// TIA Portal project "RRI" (V15.1)

(* hardware
DEVICE "S7-1200 station_1"  S7-1200 Station
   slot 0: "Rack_0"  S7-1200 Rack  Rack  V1.0
   slot 1: "PLC_1"  CPU 1215C DC/DC/DC  6ES7 215-1AG40-0XB0  V4.3
   slot 2: "AI 4xRTD_1"  SM 1231 AI4 x RTD  6ES7 231-5PD32-0XB0  V2.0
   slot 3: "DI 16/DQ 16x24VDC_1"  6ES7 223-1BL32-0XB0  V2.0
DEVICE "GSD device_2"  GSD.Device.PN
   slot 0: "Rack"  Rack  V1.0
   slot 0: "clipx_M5"  0.25 ms, 6 slots  BMxx
      slot 0: "0.25 ms, 6 slots"  0.25 ms, 6 slots
      slot 1: "PN-IO"  PN-IO
         slot 1: "Port 1"  Port 1
         slot 2: "Port 2"  Port 2
   slot 1: "Max value_1"  Max value
      slot 0: "max value (REAL)"  max value (REAL)
   slot 2: "Min value_1"  Min value
      slot 0: "min value (REAL)"  min value (REAL)
DEVICE "GSD device_1"  GSD.Device.PN
   slot 0: "Rack"  Rack  V1.0
   slot 0: "ek9300-16"  EK9300 V2.3  EK9300  V1.00
      slot 0: "EK9300 V2.3_1"  EK9300 V2.3
      slot 1: "EK9300 V2.3"  EK9300 V2.3
         slot 1: "Port 1"  Port 1
         slot 2: "Port 2"  Port 2
   slot 1: "Standard"  Standard
   slot 1: "EL3068_1"  EL3068  EL3068
      slot 0: "ModuleAccessPoint"  ModuleAccessPoint
   slot 1: "Standard"  Standard
DEVICE "GSD device_3"  GSD.Device.PN
   slot 0: "Rack"  Rack  V1.0
   slot 0: "clipx_M1"  0.25 ms, 6 slots  BMxx
      slot 0: "0.25 ms, 6 slots"  0.25 ms, 6 slots
      slot 1: "PN-IO"  PN-IO
         slot 1: "Port 1"  Port 1
         slot 2: "Port 2"  Port 2
   slot 1: "Max value_1"  Max value
      slot 0: "max value (REAL)"  max value (REAL)
   slot 2: "Min value_1"  Min value
      slot 0: "min value (REAL)"  min value (REAL)
   slot 3: "Max value_2"  Max value
      slot 0: "max value (REAL)"  max value (REAL)
   slot 4: "Min value_2"  Min value
      slot 0: "min value (REAL)"  min value (REAL)
DEVICE "GSD device_4"  GSD.Device.PN
   slot 0: "Rack"  Rack  V1.0
   slot 0: "clipx_M2"  0.25 ms, 6 slots  BMxx
      slot 0: "0.25 ms, 6 slots"  0.25 ms, 6 slots
      slot 1: "PN-IO"  PN-IO
         slot 1: "Port 1"  Port 1
         slot 2: "Port 2"  Port 2
   slot 1: "Max value_1"  Max value
      slot 0: "max value (REAL)"  max value (REAL)
   slot 2: "Min value_1"  Min value
      slot 0: "min value (REAL)"  min value (REAL)
DEVICE "GSD device_5"  GSD.Device.PN
   slot 0: "Rack"  Rack  V1.0
   slot 0: "clipx_M3"  0.25 ms, 6 slots  BMxx
      slot 0: "0.25 ms, 6 slots"  0.25 ms, 6 slots
      slot 1: "PN-IO"  PN-IO
         slot 1: "Port 1"  Port 1
         slot 2: "Port 2"  Port 2
   slot 1: "Max value_1"  Max value
      slot 0: "max value (REAL)"  max value (REAL)
   slot 2: "Min value_1"  Min value
      slot 0: "min value (REAL)"  min value (REAL)
DEVICE "GSD device_6"  GSD.Device.PN
   slot 0: "Rack"  Rack  V1.0
   slot 0: "clipx_M4"  0.25 ms, 6 slots  BMxx
      slot 0: "0.25 ms, 6 slots"  0.25 ms, 6 slots
      slot 1: "PN-IO"  PN-IO
         slot 1: "Port 1"  Port 1
         slot 2: "Port 2"  Port 2
   slot 1: "Max value_1"  Max value
      slot 0: "max value (REAL)"  max value (REAL)
   slot 2: "Min value_1"  Min value
      slot 0: "min value (REAL)"  min value (REAL)
*)

// ===== PLC "PLC_1"  CPU 1215C DC/DC/DC =====

VAR_GLOBAL   // PLC tag table "Default tag table"
   "System_Byte" AT %MB1 : Byte;
   "FirstScan" AT %M1.0 : Bool;
   "DiagStatusUpdate" AT %M1.1 : Bool;
   "AlwaysTRUE" AT %M1.2 : Bool;
   "AlwaysFALSE" AT %M1.3 : Bool;
   "Clock_Byte" AT %MB0 : Byte;
   "Clock_10Hz" AT %M0.0 : Bool;
   "Clock_5Hz" AT %M0.1 : Bool;
   "Clock_2.5Hz" AT %M0.2 : Bool;
   "Clock_2Hz" AT %M0.3 : Bool;
   "Clock_1.25Hz" AT %M0.4 : Bool;
   "Clock_1Hz" AT %M0.5 : Bool;
   "Clock_0.625Hz" AT %M0.6 : Bool;
   "Clock_0.5Hz" AT %M0.7 : Bool;
   "reserve(4)" AT %Q0.3 : Bool;
   "i_xSystemTrigger" AT %I0.0 : Bool;
   "reserve" AT %I1.1 : Bool;
   "q_xSystemOK" AT %Q0.0 : Bool;
   "q_xM1_PWR_EN" AT %Q0.5 : Bool;   // 48V DC!
   "q_xM2_PWR_EN" AT %Q0.6 : Bool;   // 48V DC!
   "q_xM3_PWR_EN" AT %Q0.7 : Bool;   // 48V DC!
   "q_xM4_PWR_EN" AT %Q1.0 : Bool;   // 48V DC!
   "i_wRTD_ch0" AT %IW112 : Int;   // RTD CH0
   "i_wRTD_ch1" AT %IW114 : Int;   // RTD CH1
   "i_iwRTD_ch2" AT %IW116 : Int;   // RTD CH2 - okolica
   "i_wRTD_ch3" AT %IW118 : Int;   // RTC CH3
   "Tag_2" AT %M20.0 : Bool;
   "Redge" AT %M2.0 : Bool;
   "m_stevecPreklopov" AT %M2.1 : Bool;
   "xtest" AT %M2.2 : Bool;
   "i_xShapeSensor2" AT %I1.5 : Bool;   // Sape of strip
   "Tag_3" AT %I68.0 : Bool;
   "reserve(5)" AT %Q0.4 : Bool;
   "reserve(2)" AT %Q0.1 : Bool;
   "reserve(3)" AT %Q0.2 : Bool;
   "i_xEncoderA" AT %I0.1 : Bool;
   "i_xEncoderB" AT %I0.2 : Bool;
   "i_xEncoderZ" AT %I0.3 : Bool;
   "i_xEgasiPWR_48V_M1" AT %I0.4 : Bool;
   "i_xEgasiPWR_48V_M2" AT %I0.5 : Bool;
   "i_xEgasiPWR_48V_M3" AT %I0.6 : Bool;
   "i_xEgasiPWR_48V_M4" AT %I0.7 : Bool;
   "i_xEgasiPWR_48V_M5" AT %I1.0 : Bool;
   "i_xDoubleFeed" AT %I1.2 : Bool;
   "i_xSmallFeed" AT %I1.3 : Bool;
   "i_xShapeSensor1" AT %I1.4 : Bool;   // Shape of strip
   "i_xM1inPOS1" AT %I16.0 : Bool;
   "i_xM1nPOS2" AT %I16.1 : Bool;
   "i_xM1isHommed" AT %I16.2 : Bool;
   "i_xM2inPOS1" AT %I16.3 : Bool;
   "i_xM2inPOS2" AT %I16.4 : Bool;
   "i_xM2isHommed" AT %I16.5 : Bool;
   "i_xM3inPOS1" AT %I16.6 : Bool;
   "i_xM3inPOS2" AT %I16.7 : Bool;
   "i_xM3isHommed" AT %I17.0 : Bool;
   "i_xM4inPOS1" AT %I17.1 : Bool;
   "i_xM4inPOS2" AT %I17.2 : Bool;
   "i_xM4isHommed" AT %I17.3 : Bool;
   "i_xM5inPOS1" AT %I17.4 : Bool;
   "i_xM5inPOS2" AT %I17.5 : Bool;
   "i_xM5isHommed" AT %I17.6 : Bool;
   "reserve(1)" AT %I17.7 : Bool;
   "q_xM5_PWR_EN" AT %Q1.1 : Bool;   // 48V DC!
   "q_xM1_goPOS1" AT %Q16.0 : Bool;
   "q_xM1_goPOS2" AT %Q16.1 : Bool;
   "q_xM1_goHOME" AT %Q16.2 : Bool;
   "q_xM2_goPOS1" AT %Q16.3 : Bool;
   "q_xM2_goPOS2" AT %Q16.4 : Bool;
   "q_xM2_goHOME" AT %Q16.5 : Bool;
   "q_xM3_goPOS1" AT %Q16.6 : Bool;
   "q_xM3_goPOS2" AT %Q16.7 : Bool;
   "q_xM3_goHOME" AT %Q17.0 : Bool;
   "q_xM4_goPOS1" AT %Q17.1 : Bool;
   "q_xM4_goPOS2" AT %Q17.2 : Bool;
   "q_xM4_goHOME" AT %Q17.3 : Bool;
   "q_xM5_goPOS1" AT %Q17.4 : Bool;
   "q_xM5_goPOS2" AT %Q17.5 : Bool;
   "q_xM5_goHOME" AT %Q17.6 : Bool;
   "6zhj" AT %Q17.7 : Bool;
   "clockmerker" AT %M3.7 : Bool;
   "xenabledemoCLock" AT %M4.0 : Bool;
   "xMotorDoublePowerON" AT %M4.1 : Bool;   // POWER FOR 2 MOTORS
   "xgoPOS1xMotorDoubleGOPOS2" AT %M4.2 : Bool;
   "xgoPOS1xMotorDoubleGOPOS1" AT %M4.3 : Bool;
   "xgoHOME" AT %M4.4 : Bool;
END_VAR

VAR_GLOBAL   // PLC tag table "TC"
   "i_wTemperatureTool1" AT %IW96 : Word;
   "i_wTemperatureTool2" AT %IW98 : Word;
   "i_wTemperatureTool3" AT %IW100 : Word;
   "i_wTemepratureTool4" AT %IW102 : Word;
   "Tag_1" AT %IW16 : Word;
   "Tag_4" AT %IW12 : Word;
   "Tag_5" AT %IW14 : Word;
END_VAR

VAR_GLOBAL   // PLC tag table "AKDs"
   "fromAKD1" AT %I80.0 : "AKD_TO_SIEMENS";
   "toAKD1" AT %Q68.0 : "SIEMENS_TO_AKD";
   "testbit" AT %M2.3 : Bool;
   "xsoftwareEnable" AT %M2.4 : Bool;
   "p_trig-FaultRelay" AT %M2.5 : Bool;
   "xDemoMode" AT %M2.6 : Bool;
   "xActuatorStatus" AT %M2.7 : Bool;
   "xActiveateDemoMode" AT %M3.0 : Bool;
   "xControlOverMachine" AT %M3.1 : Bool;
   "p_trig_trigg" AT %M3.2 : Bool;
   "tooglebit" AT %M3.3 : Bool;
   "r_eege_triger" AT %M3.4 : Bool;
   "akd_clock_trig" AT %M3.5 : Bool;
   "testbitsafety" AT %M3.6 : Bool;
END_VAR

VAR_GLOBAL   // PLC tag table "HBM"
   "i_rM5_MaxForceActuator" AT %ID72 : Real;
   "i_rM5_MinForceActuator" AT %ID76 : Real;
   "i_rM1_MaxForceAcuator" AT %ID80 : Real;
   "i_rM1_MinForceAcuator" AT %ID84 : Real;
   "i_rM2_MaxForceAcuator" AT %ID88 : Real;
   "i_rM2_MinForceAcuator" AT %ID92 : Real;
   "i_rM2_MaxForceAcuator(1)" AT %ID104 : Real;
   "i_rM2_MinForceAcuator(1)" AT %ID108 : Real;
   "i_rM3_MaxForceAcuator" AT %ID96 : Real;
   "i_rM3_MinForceAcuator" AT %ID100 : Real;
   "i_rM4_MaxForceAcuator" AT %ID120 : Real;
   "i_rM4_MinForceAcuator" AT %ID124 : Real;
END_VAR

VAR_GLOBAL   // PLC tag table "AI"
   "i_AI1_STATUS" AT %IW18 : Word;
   "i_AI1_RAW_VALUE" AT %IW20 : Word;
   "i_AI2_STATUS" AT %IW22 : Word;
   "i_AI2_RAW_VALUE" AT %IW24 : Word;
   "i_AI3_STATUS" AT %IW26 : Word;
   "i_AI3_RAW_VALUE" AT %IW28 : Word;
   "i_AI4_STATUS" AT %IW30 : Word;
   "i_AI4_RAW_VALUE" AT %IW32 : Word;
   "i_AI5_STATUS" AT %IW34 : Word;
   "i_AI5_RAW_VALUE" AT %IW36 : Word;
END_VAR

TYPE "typeMqttData"
   STRUCT
      mqttTcpParam : "typeTcpConnParam";
      mqttParam : "typeMqttParam";
      mqttUserControl : Struct
         xEnable : Bool;
         xPusblish : Bool;
         sStringToPublish : String;
         Status : "typeMqttStatus";
      END_STRUCT;
   END_STRUCT;
END_TYPE

TYPE "typeMqttStatus"
   STRUCT
      xtcpEsablished : Bool;   // True if the TCP connection has been
      xmqttEstavlished : Bool;   // True if the MQTT connection has been established
      xpublished : Bool;   // True, if the message has arrived successfully at
      xbusy : Bool;   // True, while a message or ping is sent to the
      xerror : Bool;   // True if there is an error
      istatusID : Int;   // State that cause the error
      status : DWord;   // Error message
   END_STRUCT;
END_TYPE

TYPE "typeMqttParam_1"
   STRUCT
      connectFlag : "typeMqttConnectFlags_1";
      publishFlag : "typeMqttPublishFlags_1";
      keepAlive : Word := 16#0A;
      packetIdentifier : Word := 16#10;
      clientIdentifier : String[23];   // should be PROFINET devicename
      willTopic : String[100];
      willMessage : String[100];
      userName : String[20];   // must be set, if flag "username" is true
      password : String[20];   // must be set, if flag "password" is true
      topic : String[100];
      message : Array[0..1] of String;
   END_STRUCT;
END_TYPE

TYPE "typeMqttConnectFlags_1"
   STRUCT
      cleanSession : Bool;
      will : Bool;
      willQoS_1 : Bool;   // true, if QoS = 1
      willQoS_2 : Bool;   // true, if QoS = 2
      willRetain : Bool;   // must be false, if Will flag is false
      password : Bool;   // if true, a password is required
      userName : Bool;   // if true, a username is required
   END_STRUCT;
END_TYPE

TYPE "typeTcpConnParam"
   STRUCT
      hwIdentifier : Hw_Any;
      connectionID : Conn_Ouc;
      ipAdressBroker : Array[0..3] of Byte;
      localPort : UInt;
      mqttPort : UInt := 0;
   END_STRUCT;
END_TYPE

TYPE "typeMqttParam"
   STRUCT
      connectFlag : "typeMqttConnectFlags";
      publishFlag : "typeMqttPublishFlags";
      keepAlive : Word := 16#0A;
      packetIdentifier : Word := 16#10;
      clientIdentifier : String[23];   // should be PROFINET devicename
      willTopic : String[100];
      willMessage : String[100];
      userName : String[20];   // must be set, if flag "username" is true
      password : String[20];   // must be set, if flag "password" is true
      topic : String[100];
      message : String;
   END_STRUCT;
END_TYPE

TYPE "typeMqttConnectFlags"
   STRUCT
      cleanSession : Bool;
      will : Bool;
      willQoS_1 : Bool;   // true, if QoS = 1
      willQoS_2 : Bool;   // true, if QoS = 2
      willRetain : Bool;   // must be false, if Will flag is false
      password : Bool;   // if true, a password is required
      userName : Bool;   // if true, a username is required
   END_STRUCT;
END_TYPE

TYPE "typeMqttPublishFlags"
   STRUCT
      qualityOfService : Int;   // could be 0, 1, 2
      retain : Bool;
   END_STRUCT;
END_TYPE

TYPE "typeMqttPublishFlags_1"
   STRUCT
      qualityOfService : Int;   // could be 0, 1, 2
      retain : Bool;
   END_STRUCT;
END_TYPE

TYPE "typeMqttData_1"
   STRUCT
      mqttTcpParam : "typeTcpConnParam";
      mqttParam : "typeMqttParam_1";
      mqttUserControl : Struct
         xEnable : Bool;
         xPusblish : Bool;
         sStringToPublish : String;
         Status : "typeMqttStatus";
      END_STRUCT;
   END_STRUCT;
END_TYPE

// folder: AKD

TYPE "SIEMENS_TO_AKD"
   STRUCT
      PODATKI : Struct
         oBit8_jogOn : Bool;   // b0 STW x8
         oBit9_jog2On : Bool;   // 1 STW x9
         ControlByPLC : Bool;   // 2 STW x10
         StartHomming : Bool;   // 3 STW x11
         NC_B0_b4 : Bool;   // 4 STW X12
         NC_B0_b5 : Bool;   // 5 STW x13
         NC_B0_b6 : Bool;   // 6
         NC_B0_b7 : Bool;   // 7
         SwtichOn : Bool;   // 0 / SWT x0
         NoCoastStop : Bool;   // 1 / SWT x1
         NoQuickStop : Bool;   // 2 / SWT x2
         EnableOperation : Bool;   // 3 / STW x3
         EnableRampGen : Bool;   // 4 STW x4
         UnfreezeRamp : Bool;   // 5 STW x5
         EnableSetPoint : Bool;   // 6 STW x6
         FaultAckt : Bool;   // 7 1 STW x7
         SATANW : Int;   // 0- 26 2-3
         byte4 : Byte;   // 4
         byte5 : Byte;   // 5
         MDI_TARPOS : DInt;   // 6 7 8 9
         MDI_VELOCITY : DInt;   // 10 11 12 13
         b14 : DInt;   // 14
         "15" : DInt;   // 15
         b16 : DInt;   // 16
         b17 : DInt;   // 17
         MDI_MOD : DInt;   // 18,19
      END_STRUCT;
   END_STRUCT;
END_TYPE

TYPE "AKD_TO_SIEMENS"
   STRUCT
      PODATKI_TO_SIEMENS : Struct
         ErrInRange : Bool;   // ZSW x8 - following error in range
         ContrReqByMass : Bool;   // ZSW x9
         TargetPosreached : Bool;   // ZSW x10
         HomePosSet : Bool;   // ZSW x11
         TravesingTaskAck : Bool;   // ZSW x12
         DriveStopen : Bool;   // ZSW x13
         MotionTaskActive : Bool;   // ZSW x14 - motion task active
         "i_b0.7" : Bool;   // ZSW x15 - NC
         ReadyToSwitch : Bool;   // ZSW x0
         ReadyToOperate : Bool;   // ZSW x1
         OperationENabled : Bool;   // ZSW x2
         FaultPresent : Bool;   // ZSW x3
         CoastStopNotAct : Bool;   // ZSW x4
         QuickStopNotAct : Bool;   // ZSW x5
         SwitchOnInhibiited : Bool;   // ZSW x6
         WarningPreent : Bool;   // ZSW x7
         AKTSATZ : Word;
         ZSW2 : Word;
         ActualPos : DWord;
      END_STRUCT;
   END_STRUCT;
END_TYPE

TYPE "UDT_AKD_TG400"
TITLE = UDT_AKD_TG400
VERSION : 0.1
// Matched with telegram 400 and TG400 function block.
   STRUCT
      Send : Struct
         STW1 : Int;   // Control word 1
         SATZANW : Int;   // Motion task selection
         STW2 : Int;   // Control word 2
         MDI_TARPOS : Int;   // MDI motion task target position
         MDI_TARPOS_1 : Int;   // MDI motion task target position
         MDI_VELOCITY : Int;   // MDI motion task velocity
         MDI_VELOCITY_1 : Int;   // MDI motion task velocity
         MDI_ACC : Int;   // MDI motion task acceleration
         MDI_DEC : Int;   // MDI motion task deceleration
         MDI_MOD : Int;   // MDI motion task control word
         HOME_DIST : Int;   // Home distance
         HOME_DIST_1 : Int;   // Home distance
         IDT_DATAITEM_I_12 : Int;   // Process data word input 13
         IDT_DATAITEM_I_13 : Int;   // Process data word input 14
         IDT_DATAITEM_I_14 : Int;   // Process data word input 15
         IDT_DATAITEM_I_15 : Int;   // Process data word input 16
      END_STRUCT;
      Receive : Struct
         ZSW1 : Int;   // Status word 1
         AKTSATZ : Int;   // Actual motion task selection
         ZSW2 : Int;   // Status word 2
         XIST_A : Int;   // Actual position
         XIST_A_1 : Int;   // Actual position
         NIST_A : Int;   // Actual velocity
         ITIST_GLATT : Int;   // Actual current
         IDT_DATAITEM_O_7 : Int;   // Process data word output 8
         IDT_DATAITEM_O_8 : Int;   // Process data word output 9
         IDT_DATAITEM_O_9 : Int;   // Process data word output 10
         IDT_DATAITEM_O_10 : Int;   // Process data word output 11
         IDT_DATAITEM_O_11 : Int;   // Process data word output 12
         IDT_DATAITEM_O_12 : Int;   // Process data word output 13
         IDT_DATAITEM_O_13 : Int;   // Process data word output 14
         IDT_DATAITEM_O_14 : Int;   // Process data word output 15
         IDT_DATAITEM_O_15 : Int;   // Process data word output 16
      END_STRUCT;
   END_STRUCT;
END_TYPE

// folder: AKD/PNU

TYPE "AKD_FROM_PNU"
   STRUCT
      xActive : Bool;
      xDone : Bool;
      xError : Bool;
      dStatus : DInt;
   END_STRUCT;
END_TYPE

TYPE "AKD_TO_PNU"
   STRUCT
      iID : Hw_Io;   // HW ID of a AKD
      xStartReq : Bool;   // start request
      xReqType : Bool;   // 0-read, 1-write
      wFormat : Word := W#16#42;   // 16#41 - byte, 16#42 -. word, 16#43 - dword
      iPNUnumber : Int;
      iPNUsubindex : Int;
      data : DInt;
      cmd : Struct
         xStartRead : Bool;
         xStartWrite : Bool;
      END_STRUCT;
      cfg : Struct
         xempty : Bool;
      END_STRUCT;
   END_STRUCT;
END_TYPE

TYPE "PNU_DATA"
   STRUCT
      to_PNU : "AKD_TO_PNU";
      From_PNU : "AKD_FROM_PNU";
   END_STRUCT;
END_TYPE

// folder: EGASI

TYPE "RRI_izdelki"
   STRUCT
      NazivniPodatki : Struct
         SifraIzdelka : Int;
         st_pomikov : Int;
         st_celic : Int;
         st_vrst : Int;
         CILINDRI : Struct
            MOTOR1 : Array[0..20] of Bool;
            MOTOR2 : Array[0..20] of Bool;
            MOTOR3 : Array[0..20] of Bool;
            MOTOR4 : Array[0..20] of Bool;
            MOTOR5 : Array[0..20] of Bool;
            MOTOR6 : Array[0..20] of Bool;
         END_STRUCT;
      END_STRUCT;
      TrenutniPodatki : Struct
         trenutni_pomik : Int;
      END_STRUCT;
      Oblika : Struct
         s1 : Array[0..20] of Bool;
         s2 : Array[0..20] of Bool;
      END_STRUCT;
   END_STRUCT;
END_TYPE

TYPE "EGASI_MOTOR_CONTROL"
   STRUCT
      fromMOTOR : Struct
         xInPOS1 : Bool;
         xinPOS2 : Bool;
         xisHOMMED : Bool;
         wRawTempValue : Word;
         rScaledTempValue : Real;
         rRawCurrentMAXValue : Real;
         rRawCurrentMINvalue : Real;
         xPowerStatus : Bool;   // is Power ON/OFF?
      END_STRUCT;
      toMOTOR : Struct
         xPWR_EN : Bool;
         xGoPOS1 : Bool;
         xGoPOS2 : Bool;
         xGoHOME : Bool;
      END_STRUCT;
      Errors : Struct
         POS1_POS2_ERR : Bool;
         FUSE_ERR : Bool;
         POS1_notAccesible : Bool;
         POS2_notAccessible : Bool;
      END_STRUCT;
      Control : Struct
         xGoPOS1 : Bool;
         xGoPOS2 : Bool;
         xGoHome : Bool;
         xPWR_en : Bool;
         xDemoClock : Bool;
         xAutomaticMachineMode : Bool;
      END_STRUCT;
   END_STRUCT;
END_TYPE

// folder: Node-Red

TYPE "UDT_MotorDataStatus"
   STRUCT
      xinPOS1 : Bool;
      xinPOS2 : Bool;
      xisHOMMED : Bool;
      xinError : Bool;
      xFuseError : Bool;
      xPOS1Error : Bool;
      xPOS2Error : Bool;
      xPWRstatus : Bool;
      rTemperature : Real;
      rMaxForce : Real;
      rMinForce : Real;
   END_STRUCT;
END_TYPE

TYPE "UDT_MotorControl"
   STRUCT
      xGoPos1 : Bool;
      xGoPos2 : Bool;
      xGOHOME : Bool;
      xHW_reset : Bool;
   END_STRUCT;
END_TYPE

// folder: (top level)

DATA_BLOCK "FB_TcConvert_DB_TC3_TempOkolice"   // DB2
{ S7_Optimized_Access := 'TRUE' }
VERSION : 0.1
// stored: InstanceOfName FB_TcConvert
"FB_TcConvert"
BEGIN
END_DATA_BLOCK

DATA_BLOCK "DB_GlobalData"   // DB3
{ S7_Optimized_Access := 'TRUE' }
VERSION : 0.1
   VAR RETAIN
      Thermocouplers : Struct
         Thermocoupler1_tempOrodja1 : Real := 4943.8;
         Thermocoupler1_tempOrodja2 : Real := 1060.6;
         Thermocoupler1_tempOrodja3_temperaturaOkolice : Real := 4944.1;
         Thermocoupler1_tempOrodja4 : Real := 5366.7;
      END_STRUCT;
   END_VAR
   VAR
      RTDs : Struct
         RTD1 : Struct
            ch0 : Real := -1.0;
            ch1 : Real := -1.0;
            ch2 : Real := 27.5;
            ch3 : Real := -1.0;
         END_STRUCT;
      END_STRUCT;
   END_VAR
   VAR RETAIN
      AKD : Struct
         AKD1 : Struct
            xServoRelayOn : Bool := FALSE;
            xServoProfinetOn : Bool := FALSE;
            sFaultRelay : Bool := FALSE;
            xErrorReset : Bool := FALSE;
            xStartHomming : Bool := FALSE;
            xServoGo : Bool := FALSE;
            wJobNumber : Word := 16#0000;
            wNewJobNumber : Word := 16#0000;
            Status : Struct
               status : Byte := 16#0A;
            END_STRUCT;
            resistance : Real := 0.0;
            calculatedTemp : Real := -319.85;
         END_STRUCT;
      END_STRUCT;
      Prezracevanje : Struct
         xEnableFaninManual : Bool := FALSE;
      END_STRUCT;
      Stiskalnica : Struct
         iPresaHitrost : Int := 0;
         xPresaON : Int := 0;
         uPresaStevec : UDInt := 0;
      END_STRUCT;
      PartManagmenent : Struct
         PartsToMade : "RRI_izdelki";
         LastPart : "RRI_izdelki";
         PartRecept : "RRI_izdelki";
         PartNumberForProduction : String := '39900-2';
         LastPartForProduction : String := '39900-2';
         xChangePartInProgres : Bool := FALSE;
         uiChangePartCounter : UDInt := 0;
         Trenutni_pomik : Int := 7;
         xLerningButton : Bool;
         xManualMoveLerningData : Bool;
         xAutoamtocMoveLerningData : Bool;
         xMerkers : Array[0..1] of Bool;
      END_STRUCT;
   END_VAR
BEGIN
   PartManagmenent.PartsToMade.NazivniPodatki.SifraIzdelka := 0;
   PartManagmenent.PartsToMade.NazivniPodatki.st_pomikov := 8;
   PartManagmenent.PartsToMade.NazivniPodatki.st_celic := 8;
   PartManagmenent.PartsToMade.NazivniPodatki.st_vrst := 2;
   PartManagmenent.PartsToMade.NazivniPodatki.CILINDRI.MOTOR1[1] := FALSE;
   PartManagmenent.PartsToMade.NazivniPodatki.CILINDRI.MOTOR1[2] := FALSE;
   PartManagmenent.PartsToMade.NazivniPodatki.CILINDRI.MOTOR1[3] := TRUE;
   PartManagmenent.PartsToMade.NazivniPodatki.CILINDRI.MOTOR1[4] := FALSE;
   PartManagmenent.PartsToMade.NazivniPodatki.CILINDRI.MOTOR1[5] := FALSE;
   PartManagmenent.PartsToMade.NazivniPodatki.CILINDRI.MOTOR1[6] := FALSE;
   PartManagmenent.PartsToMade.NazivniPodatki.CILINDRI.MOTOR1[7] := FALSE;
   PartManagmenent.PartsToMade.NazivniPodatki.CILINDRI.MOTOR1[8] := FALSE;
   PartManagmenent.PartsToMade.NazivniPodatki.CILINDRI.MOTOR1[9] := FALSE;
   PartManagmenent.PartsToMade.NazivniPodatki.CILINDRI.MOTOR1[10] := FALSE;
   PartManagmenent.PartsToMade.NazivniPodatki.CILINDRI.MOTOR1[11] := FALSE;
   PartManagmenent.PartsToMade.NazivniPodatki.CILINDRI.MOTOR1[12] := FALSE;
   PartManagmenent.PartsToMade.NazivniPodatki.CILINDRI.MOTOR1[13] := FALSE;
   PartManagmenent.PartsToMade.NazivniPodatki.CILINDRI.MOTOR1[14] := FALSE;
   PartManagmenent.PartsToMade.NazivniPodatki.CILINDRI.MOTOR1[15] := FALSE;
   PartManagmenent.PartsToMade.NazivniPodatki.CILINDRI.MOTOR1[16] := FALSE;
   PartManagmenent.PartsToMade.NazivniPodatki.CILINDRI.MOTOR1[17] := FALSE;
   PartManagmenent.PartsToMade.NazivniPodatki.CILINDRI.MOTOR1[18] := FALSE;
   PartManagmenent.PartsToMade.NazivniPodatki.CILINDRI.MOTOR1[19] := FALSE;
   PartManagmenent.PartsToMade.NazivniPodatki.CILINDRI.MOTOR1[20] := FALSE;
   PartManagmenent.PartsToMade.NazivniPodatki.CILINDRI.MOTOR2[1] := FALSE;
   PartManagmenent.PartsToMade.NazivniPodatki.CILINDRI.MOTOR2[2] := FALSE;
   PartManagmenent.PartsToMade.NazivniPodatki.CILINDRI.MOTOR2[3] := FALSE;
   PartManagmenent.PartsToMade.NazivniPodatki.CILINDRI.MOTOR2[4] := FALSE;
   PartManagmenent.PartsToMade.NazivniPodatki.CILINDRI.MOTOR2[5] := FALSE;
   PartManagmenent.PartsToMade.NazivniPodatki.CILINDRI.MOTOR2[6] := FALSE;
   PartManagmenent.PartsToMade.NazivniPodatki.CILINDRI.MOTOR2[7] := FALSE;
   PartManagmenent.PartsToMade.NazivniPodatki.CILINDRI.MOTOR2[8] := FALSE;
   PartManagmenent.PartsToMade.NazivniPodatki.CILINDRI.MOTOR2[9] := FALSE;
   PartManagmenent.PartsToMade.NazivniPodatki.CILINDRI.MOTOR2[10] := FALSE;
   PartManagmenent.PartsToMade.NazivniPodatki.CILINDRI.MOTOR2[11] := FALSE;
   PartManagmenent.PartsToMade.NazivniPodatki.CILINDRI.MOTOR2[12] := FALSE;
   PartManagmenent.PartsToMade.NazivniPodatki.CILINDRI.MOTOR2[13] := FALSE;
   PartManagmenent.PartsToMade.NazivniPodatki.CILINDRI.MOTOR2[14] := FALSE;
   PartManagmenent.PartsToMade.NazivniPodatki.CILINDRI.MOTOR2[15] := FALSE;
   PartManagmenent.PartsToMade.NazivniPodatki.CILINDRI.MOTOR2[16] := FALSE;
   PartManagmenent.PartsToMade.NazivniPodatki.CILINDRI.MOTOR2[17] := FALSE;
   PartManagmenent.PartsToMade.NazivniPodatki.CILINDRI.MOTOR2[18] := FALSE;
   PartManagmenent.PartsToMade.NazivniPodatki.CILINDRI.MOTOR2[19] := FALSE;
   PartManagmenent.PartsToMade.NazivniPodatki.CILINDRI.MOTOR2[20] := FALSE;
   PartManagmenent.PartsToMade.NazivniPodatki.CILINDRI.MOTOR3[1] := FALSE;
   PartManagmenent.PartsToMade.NazivniPodatki.CILINDRI.MOTOR3[2] := FALSE;
   PartManagmenent.PartsToMade.NazivniPodatki.CILINDRI.MOTOR3[3] := FALSE;
   PartManagmenent.PartsToMade.NazivniPodatki.CILINDRI.MOTOR3[4] := FALSE;
   PartManagmenent.PartsToMade.NazivniPodatki.CILINDRI.MOTOR3[5] := FALSE;
   PartManagmenent.PartsToMade.NazivniPodatki.CILINDRI.MOTOR3[6] := FALSE;
   PartManagmenent.PartsToMade.NazivniPodatki.CILINDRI.MOTOR3[7] := FALSE;
   PartManagmenent.PartsToMade.NazivniPodatki.CILINDRI.MOTOR3[8] := FALSE;
   PartManagmenent.PartsToMade.NazivniPodatki.CILINDRI.MOTOR3[9] := FALSE;
   PartManagmenent.PartsToMade.NazivniPodatki.CILINDRI.MOTOR3[10] := FALSE;
   PartManagmenent.PartsToMade.NazivniPodatki.CILINDRI.MOTOR3[11] := FALSE;
   PartManagmenent.PartsToMade.NazivniPodatki.CILINDRI.MOTOR3[12] := FALSE;
   PartManagmenent.PartsToMade.NazivniPodatki.CILINDRI.MOTOR3[13] := FALSE;
   PartManagmenent.PartsToMade.NazivniPodatki.CILINDRI.MOTOR3[14] := FALSE;
   PartManagmenent.PartsToMade.NazivniPodatki.CILINDRI.MOTOR3[15] := FALSE;
   PartManagmenent.PartsToMade.NazivniPodatki.CILINDRI.MOTOR3[16] := FALSE;
   PartManagmenent.PartsToMade.NazivniPodatki.CILINDRI.MOTOR3[17] := FALSE;
   PartManagmenent.PartsToMade.NazivniPodatki.CILINDRI.MOTOR3[18] := FALSE;
   PartManagmenent.PartsToMade.NazivniPodatki.CILINDRI.MOTOR3[19] := FALSE;
   PartManagmenent.PartsToMade.NazivniPodatki.CILINDRI.MOTOR3[20] := FALSE;
   PartManagmenent.PartsToMade.NazivniPodatki.CILINDRI.MOTOR4[1] := FALSE;
   PartManagmenent.PartsToMade.NazivniPodatki.CILINDRI.MOTOR4[2] := FALSE;
   PartManagmenent.PartsToMade.NazivniPodatki.CILINDRI.MOTOR4[3] := FALSE;
   PartManagmenent.PartsToMade.NazivniPodatki.CILINDRI.MOTOR4[4] := FALSE;
   PartManagmenent.PartsToMade.NazivniPodatki.CILINDRI.MOTOR4[5] := FALSE;
   PartManagmenent.PartsToMade.NazivniPodatki.CILINDRI.MOTOR4[6] := FALSE;
   PartManagmenent.PartsToMade.NazivniPodatki.CILINDRI.MOTOR4[7] := FALSE;
   PartManagmenent.PartsToMade.NazivniPodatki.CILINDRI.MOTOR4[8] := FALSE;
   PartManagmenent.PartsToMade.NazivniPodatki.CILINDRI.MOTOR4[9] := FALSE;
   PartManagmenent.PartsToMade.NazivniPodatki.CILINDRI.MOTOR4[10] := FALSE;
   PartManagmenent.PartsToMade.NazivniPodatki.CILINDRI.MOTOR4[11] := FALSE;
   PartManagmenent.PartsToMade.NazivniPodatki.CILINDRI.MOTOR4[12] := FALSE;
   PartManagmenent.PartsToMade.NazivniPodatki.CILINDRI.MOTOR4[13] := FALSE;
   PartManagmenent.PartsToMade.NazivniPodatki.CILINDRI.MOTOR4[14] := FALSE;
   PartManagmenent.PartsToMade.NazivniPodatki.CILINDRI.MOTOR4[15] := FALSE;
   PartManagmenent.PartsToMade.NazivniPodatki.CILINDRI.MOTOR4[16] := FALSE;
   PartManagmenent.PartsToMade.NazivniPodatki.CILINDRI.MOTOR4[17] := FALSE;
   PartManagmenent.PartsToMade.NazivniPodatki.CILINDRI.MOTOR4[18] := FALSE;
   PartManagmenent.PartsToMade.NazivniPodatki.CILINDRI.MOTOR4[19] := FALSE;
   PartManagmenent.PartsToMade.NazivniPodatki.CILINDRI.MOTOR4[20] := FALSE;
   PartManagmenent.PartsToMade.NazivniPodatki.CILINDRI.MOTOR5[1] := FALSE;
   PartManagmenent.PartsToMade.NazivniPodatki.CILINDRI.MOTOR5[2] := FALSE;
   PartManagmenent.PartsToMade.NazivniPodatki.CILINDRI.MOTOR5[3] := FALSE;
   PartManagmenent.PartsToMade.NazivniPodatki.CILINDRI.MOTOR5[4] := FALSE;
   PartManagmenent.PartsToMade.NazivniPodatki.CILINDRI.MOTOR5[5] := FALSE;
   PartManagmenent.PartsToMade.NazivniPodatki.CILINDRI.MOTOR5[6] := FALSE;
   PartManagmenent.PartsToMade.NazivniPodatki.CILINDRI.MOTOR5[7] := FALSE;
   PartManagmenent.PartsToMade.NazivniPodatki.CILINDRI.MOTOR5[8] := FALSE;
   PartManagmenent.PartsToMade.NazivniPodatki.CILINDRI.MOTOR5[9] := FALSE;
   PartManagmenent.PartsToMade.NazivniPodatki.CILINDRI.MOTOR5[10] := FALSE;
   PartManagmenent.PartsToMade.NazivniPodatki.CILINDRI.MOTOR5[11] := FALSE;
   PartManagmenent.PartsToMade.NazivniPodatki.CILINDRI.MOTOR5[12] := FALSE;
   PartManagmenent.PartsToMade.NazivniPodatki.CILINDRI.MOTOR5[13] := FALSE;
   PartManagmenent.PartsToMade.NazivniPodatki.CILINDRI.MOTOR5[14] := FALSE;
   PartManagmenent.PartsToMade.NazivniPodatki.CILINDRI.MOTOR5[15] := FALSE;
   PartManagmenent.PartsToMade.NazivniPodatki.CILINDRI.MOTOR5[16] := FALSE;
   PartManagmenent.PartsToMade.NazivniPodatki.CILINDRI.MOTOR5[17] := FALSE;
   PartManagmenent.PartsToMade.NazivniPodatki.CILINDRI.MOTOR5[18] := FALSE;
   PartManagmenent.PartsToMade.NazivniPodatki.CILINDRI.MOTOR5[19] := FALSE;
   PartManagmenent.PartsToMade.NazivniPodatki.CILINDRI.MOTOR5[20] := FALSE;
   PartManagmenent.PartsToMade.NazivniPodatki.CILINDRI.MOTOR6[1] := FALSE;
   PartManagmenent.PartsToMade.NazivniPodatki.CILINDRI.MOTOR6[2] := FALSE;
   PartManagmenent.PartsToMade.NazivniPodatki.CILINDRI.MOTOR6[3] := FALSE;
   PartManagmenent.PartsToMade.NazivniPodatki.CILINDRI.MOTOR6[4] := FALSE;
   PartManagmenent.PartsToMade.NazivniPodatki.CILINDRI.MOTOR6[5] := FALSE;
   PartManagmenent.PartsToMade.NazivniPodatki.CILINDRI.MOTOR6[6] := FALSE;
   PartManagmenent.PartsToMade.NazivniPodatki.CILINDRI.MOTOR6[7] := FALSE;
   PartManagmenent.PartsToMade.NazivniPodatki.CILINDRI.MOTOR6[8] := FALSE;
   PartManagmenent.PartsToMade.NazivniPodatki.CILINDRI.MOTOR6[9] := FALSE;
   PartManagmenent.PartsToMade.NazivniPodatki.CILINDRI.MOTOR6[10] := FALSE;
   PartManagmenent.PartsToMade.NazivniPodatki.CILINDRI.MOTOR6[11] := FALSE;
   PartManagmenent.PartsToMade.NazivniPodatki.CILINDRI.MOTOR6[12] := FALSE;
   PartManagmenent.PartsToMade.NazivniPodatki.CILINDRI.MOTOR6[13] := FALSE;
   PartManagmenent.PartsToMade.NazivniPodatki.CILINDRI.MOTOR6[14] := FALSE;
   PartManagmenent.PartsToMade.NazivniPodatki.CILINDRI.MOTOR6[15] := FALSE;
   PartManagmenent.PartsToMade.NazivniPodatki.CILINDRI.MOTOR6[16] := FALSE;
   PartManagmenent.PartsToMade.NazivniPodatki.CILINDRI.MOTOR6[17] := FALSE;
   PartManagmenent.PartsToMade.NazivniPodatki.CILINDRI.MOTOR6[18] := FALSE;
   PartManagmenent.PartsToMade.NazivniPodatki.CILINDRI.MOTOR6[19] := FALSE;
   PartManagmenent.PartsToMade.NazivniPodatki.CILINDRI.MOTOR6[20] := FALSE;
   PartManagmenent.PartsToMade.TrenutniPodatki.trenutni_pomik := 3350;
   PartManagmenent.PartsToMade.Oblika.s1[0] := FALSE;
   PartManagmenent.PartsToMade.Oblika.s1[1] := FALSE;
   PartManagmenent.PartsToMade.Oblika.s1[2] := FALSE;
   PartManagmenent.PartsToMade.Oblika.s1[3] := FALSE;
   PartManagmenent.PartsToMade.Oblika.s1[4] := FALSE;
   PartManagmenent.PartsToMade.Oblika.s1[5] := FALSE;
   PartManagmenent.PartsToMade.Oblika.s1[6] := FALSE;
   PartManagmenent.PartsToMade.Oblika.s1[7] := FALSE;
   PartManagmenent.PartsToMade.Oblika.s1[8] := FALSE;
   PartManagmenent.PartsToMade.Oblika.s1[9] := FALSE;
   PartManagmenent.PartsToMade.Oblika.s1[10] := FALSE;
   PartManagmenent.PartsToMade.Oblika.s1[11] := FALSE;
   PartManagmenent.PartsToMade.Oblika.s1[12] := FALSE;
   PartManagmenent.PartsToMade.Oblika.s1[13] := FALSE;
   PartManagmenent.PartsToMade.Oblika.s1[14] := FALSE;
   PartManagmenent.PartsToMade.Oblika.s1[15] := FALSE;
   PartManagmenent.PartsToMade.Oblika.s1[16] := FALSE;
   PartManagmenent.PartsToMade.Oblika.s1[17] := FALSE;
   PartManagmenent.PartsToMade.Oblika.s1[18] := FALSE;
   PartManagmenent.PartsToMade.Oblika.s1[19] := FALSE;
   PartManagmenent.PartsToMade.Oblika.s1[20] := FALSE;
   PartManagmenent.PartsToMade.Oblika.s2[0] := FALSE;
   PartManagmenent.PartsToMade.Oblika.s2[1] := FALSE;
   PartManagmenent.PartsToMade.Oblika.s2[2] := FALSE;
   PartManagmenent.PartsToMade.Oblika.s2[3] := FALSE;
   PartManagmenent.PartsToMade.Oblika.s2[4] := FALSE;
   PartManagmenent.PartsToMade.Oblika.s2[5] := FALSE;
   PartManagmenent.PartsToMade.Oblika.s2[6] := FALSE;
   PartManagmenent.PartsToMade.Oblika.s2[7] := FALSE;
   PartManagmenent.PartsToMade.Oblika.s2[8] := FALSE;
   PartManagmenent.PartsToMade.Oblika.s2[9] := FALSE;
   PartManagmenent.PartsToMade.Oblika.s2[10] := FALSE;
   PartManagmenent.PartsToMade.Oblika.s2[11] := FALSE;
   PartManagmenent.PartsToMade.Oblika.s2[12] := FALSE;
   PartManagmenent.PartsToMade.Oblika.s2[13] := FALSE;
   PartManagmenent.PartsToMade.Oblika.s2[14] := FALSE;
   PartManagmenent.PartsToMade.Oblika.s2[15] := FALSE;
   PartManagmenent.PartsToMade.Oblika.s2[16] := FALSE;
   PartManagmenent.PartsToMade.Oblika.s2[17] := FALSE;
   PartManagmenent.PartsToMade.Oblika.s2[18] := FALSE;
   PartManagmenent.PartsToMade.Oblika.s2[19] := FALSE;
   PartManagmenent.PartsToMade.Oblika.s2[20] := FALSE;
   PartManagmenent.LastPart.NazivniPodatki.SifraIzdelka := 0;
   PartManagmenent.LastPart.NazivniPodatki.st_pomikov := 4;
   PartManagmenent.LastPart.NazivniPodatki.st_celic := 4;
   PartManagmenent.LastPart.NazivniPodatki.st_vrst := 2;
   PartManagmenent.LastPart.NazivniPodatki.CILINDRI.MOTOR1[1] := FALSE;
   PartManagmenent.LastPart.NazivniPodatki.CILINDRI.MOTOR1[2] := TRUE;
   PartManagmenent.LastPart.NazivniPodatki.CILINDRI.MOTOR1[3] := FALSE;
   PartManagmenent.LastPart.NazivniPodatki.CILINDRI.MOTOR1[4] := FALSE;
   PartManagmenent.LastPart.NazivniPodatki.CILINDRI.MOTOR1[5] := FALSE;
   PartManagmenent.LastPart.NazivniPodatki.CILINDRI.MOTOR1[6] := FALSE;
   PartManagmenent.LastPart.NazivniPodatki.CILINDRI.MOTOR1[7] := FALSE;
   PartManagmenent.LastPart.NazivniPodatki.CILINDRI.MOTOR1[8] := FALSE;
   PartManagmenent.LastPart.NazivniPodatki.CILINDRI.MOTOR1[9] := FALSE;
   PartManagmenent.LastPart.NazivniPodatki.CILINDRI.MOTOR1[10] := FALSE;
   PartManagmenent.LastPart.NazivniPodatki.CILINDRI.MOTOR1[11] := FALSE;
   PartManagmenent.LastPart.NazivniPodatki.CILINDRI.MOTOR1[12] := FALSE;
   PartManagmenent.LastPart.NazivniPodatki.CILINDRI.MOTOR1[13] := FALSE;
   PartManagmenent.LastPart.NazivniPodatki.CILINDRI.MOTOR1[14] := FALSE;
   PartManagmenent.LastPart.NazivniPodatki.CILINDRI.MOTOR1[15] := FALSE;
   PartManagmenent.LastPart.NazivniPodatki.CILINDRI.MOTOR1[16] := FALSE;
   PartManagmenent.LastPart.NazivniPodatki.CILINDRI.MOTOR1[17] := FALSE;
   PartManagmenent.LastPart.NazivniPodatki.CILINDRI.MOTOR1[18] := FALSE;
   PartManagmenent.LastPart.NazivniPodatki.CILINDRI.MOTOR1[19] := FALSE;
   PartManagmenent.LastPart.NazivniPodatki.CILINDRI.MOTOR1[20] := FALSE;
   PartManagmenent.LastPart.NazivniPodatki.CILINDRI.MOTOR2[1] := FALSE;
   PartManagmenent.LastPart.NazivniPodatki.CILINDRI.MOTOR2[2] := FALSE;
   PartManagmenent.LastPart.NazivniPodatki.CILINDRI.MOTOR2[3] := FALSE;
   PartManagmenent.LastPart.NazivniPodatki.CILINDRI.MOTOR2[4] := FALSE;
   PartManagmenent.LastPart.NazivniPodatki.CILINDRI.MOTOR2[5] := FALSE;
   PartManagmenent.LastPart.NazivniPodatki.CILINDRI.MOTOR2[6] := FALSE;
   PartManagmenent.LastPart.NazivniPodatki.CILINDRI.MOTOR2[7] := FALSE;
   PartManagmenent.LastPart.NazivniPodatki.CILINDRI.MOTOR2[8] := FALSE;
   PartManagmenent.LastPart.NazivniPodatki.CILINDRI.MOTOR2[9] := FALSE;
   PartManagmenent.LastPart.NazivniPodatki.CILINDRI.MOTOR2[10] := FALSE;
   PartManagmenent.LastPart.NazivniPodatki.CILINDRI.MOTOR2[11] := FALSE;
   PartManagmenent.LastPart.NazivniPodatki.CILINDRI.MOTOR2[12] := FALSE;
   PartManagmenent.LastPart.NazivniPodatki.CILINDRI.MOTOR2[13] := FALSE;
   PartManagmenent.LastPart.NazivniPodatki.CILINDRI.MOTOR2[14] := FALSE;
   PartManagmenent.LastPart.NazivniPodatki.CILINDRI.MOTOR2[15] := FALSE;
   PartManagmenent.LastPart.NazivniPodatki.CILINDRI.MOTOR2[16] := FALSE;
   PartManagmenent.LastPart.NazivniPodatki.CILINDRI.MOTOR2[17] := FALSE;
   PartManagmenent.LastPart.NazivniPodatki.CILINDRI.MOTOR2[18] := FALSE;
   PartManagmenent.LastPart.NazivniPodatki.CILINDRI.MOTOR2[19] := FALSE;
   PartManagmenent.LastPart.NazivniPodatki.CILINDRI.MOTOR2[20] := FALSE;
   PartManagmenent.LastPart.NazivniPodatki.CILINDRI.MOTOR3[1] := FALSE;
   PartManagmenent.LastPart.NazivniPodatki.CILINDRI.MOTOR3[2] := FALSE;
   PartManagmenent.LastPart.NazivniPodatki.CILINDRI.MOTOR3[3] := FALSE;
   PartManagmenent.LastPart.NazivniPodatki.CILINDRI.MOTOR3[4] := FALSE;
   PartManagmenent.LastPart.NazivniPodatki.CILINDRI.MOTOR3[5] := FALSE;
   PartManagmenent.LastPart.NazivniPodatki.CILINDRI.MOTOR3[6] := FALSE;
   PartManagmenent.LastPart.NazivniPodatki.CILINDRI.MOTOR3[7] := FALSE;
   PartManagmenent.LastPart.NazivniPodatki.CILINDRI.MOTOR3[8] := FALSE;
   PartManagmenent.LastPart.NazivniPodatki.CILINDRI.MOTOR3[9] := FALSE;
   PartManagmenent.LastPart.NazivniPodatki.CILINDRI.MOTOR3[10] := FALSE;
   PartManagmenent.LastPart.NazivniPodatki.CILINDRI.MOTOR3[11] := FALSE;
   PartManagmenent.LastPart.NazivniPodatki.CILINDRI.MOTOR3[12] := FALSE;
   PartManagmenent.LastPart.NazivniPodatki.CILINDRI.MOTOR3[13] := FALSE;
   PartManagmenent.LastPart.NazivniPodatki.CILINDRI.MOTOR3[14] := FALSE;
   PartManagmenent.LastPart.NazivniPodatki.CILINDRI.MOTOR3[15] := FALSE;
   PartManagmenent.LastPart.NazivniPodatki.CILINDRI.MOTOR3[16] := FALSE;
   PartManagmenent.LastPart.NazivniPodatki.CILINDRI.MOTOR3[17] := FALSE;
   PartManagmenent.LastPart.NazivniPodatki.CILINDRI.MOTOR3[18] := FALSE;
   PartManagmenent.LastPart.NazivniPodatki.CILINDRI.MOTOR3[19] := FALSE;
   PartManagmenent.LastPart.NazivniPodatki.CILINDRI.MOTOR3[20] := FALSE;
   PartManagmenent.LastPart.NazivniPodatki.CILINDRI.MOTOR4[1] := FALSE;
   PartManagmenent.LastPart.NazivniPodatki.CILINDRI.MOTOR4[2] := FALSE;
   PartManagmenent.LastPart.NazivniPodatki.CILINDRI.MOTOR4[3] := FALSE;
   PartManagmenent.LastPart.NazivniPodatki.CILINDRI.MOTOR4[4] := FALSE;
   PartManagmenent.LastPart.NazivniPodatki.CILINDRI.MOTOR4[5] := FALSE;
   PartManagmenent.LastPart.NazivniPodatki.CILINDRI.MOTOR4[6] := FALSE;
   PartManagmenent.LastPart.NazivniPodatki.CILINDRI.MOTOR4[7] := FALSE;
   PartManagmenent.LastPart.NazivniPodatki.CILINDRI.MOTOR4[8] := FALSE;
   PartManagmenent.LastPart.NazivniPodatki.CILINDRI.MOTOR4[9] := FALSE;
   PartManagmenent.LastPart.NazivniPodatki.CILINDRI.MOTOR4[10] := FALSE;
   PartManagmenent.LastPart.NazivniPodatki.CILINDRI.MOTOR4[11] := FALSE;
   PartManagmenent.LastPart.NazivniPodatki.CILINDRI.MOTOR4[12] := FALSE;
   PartManagmenent.LastPart.NazivniPodatki.CILINDRI.MOTOR4[13] := FALSE;
   PartManagmenent.LastPart.NazivniPodatki.CILINDRI.MOTOR4[14] := FALSE;
   PartManagmenent.LastPart.NazivniPodatki.CILINDRI.MOTOR4[15] := FALSE;
   PartManagmenent.LastPart.NazivniPodatki.CILINDRI.MOTOR4[16] := FALSE;
   PartManagmenent.LastPart.NazivniPodatki.CILINDRI.MOTOR4[17] := FALSE;
   PartManagmenent.LastPart.NazivniPodatki.CILINDRI.MOTOR4[18] := FALSE;
   PartManagmenent.LastPart.NazivniPodatki.CILINDRI.MOTOR4[19] := FALSE;
   PartManagmenent.LastPart.NazivniPodatki.CILINDRI.MOTOR4[20] := FALSE;
   PartManagmenent.LastPart.NazivniPodatki.CILINDRI.MOTOR5[1] := FALSE;
   PartManagmenent.LastPart.NazivniPodatki.CILINDRI.MOTOR5[2] := FALSE;
   PartManagmenent.LastPart.NazivniPodatki.CILINDRI.MOTOR5[3] := FALSE;
   PartManagmenent.LastPart.NazivniPodatki.CILINDRI.MOTOR5[4] := FALSE;
   PartManagmenent.LastPart.NazivniPodatki.CILINDRI.MOTOR5[5] := FALSE;
   PartManagmenent.LastPart.NazivniPodatki.CILINDRI.MOTOR5[6] := FALSE;
   PartManagmenent.LastPart.NazivniPodatki.CILINDRI.MOTOR5[7] := FALSE;
   PartManagmenent.LastPart.NazivniPodatki.CILINDRI.MOTOR5[8] := FALSE;
   PartManagmenent.LastPart.NazivniPodatki.CILINDRI.MOTOR5[9] := FALSE;
   PartManagmenent.LastPart.NazivniPodatki.CILINDRI.MOTOR5[10] := FALSE;
   PartManagmenent.LastPart.NazivniPodatki.CILINDRI.MOTOR5[11] := FALSE;
   PartManagmenent.LastPart.NazivniPodatki.CILINDRI.MOTOR5[12] := FALSE;
   PartManagmenent.LastPart.NazivniPodatki.CILINDRI.MOTOR5[13] := FALSE;
   PartManagmenent.LastPart.NazivniPodatki.CILINDRI.MOTOR5[14] := FALSE;
   PartManagmenent.LastPart.NazivniPodatki.CILINDRI.MOTOR5[15] := FALSE;
   PartManagmenent.LastPart.NazivniPodatki.CILINDRI.MOTOR5[16] := FALSE;
   PartManagmenent.LastPart.NazivniPodatki.CILINDRI.MOTOR5[17] := FALSE;
   PartManagmenent.LastPart.NazivniPodatki.CILINDRI.MOTOR5[18] := FALSE;
   PartManagmenent.LastPart.NazivniPodatki.CILINDRI.MOTOR5[19] := FALSE;
   PartManagmenent.LastPart.NazivniPodatki.CILINDRI.MOTOR5[20] := FALSE;
   PartManagmenent.LastPart.NazivniPodatki.CILINDRI.MOTOR6[1] := FALSE;
   PartManagmenent.LastPart.NazivniPodatki.CILINDRI.MOTOR6[2] := FALSE;
   PartManagmenent.LastPart.NazivniPodatki.CILINDRI.MOTOR6[3] := FALSE;
   PartManagmenent.LastPart.NazivniPodatki.CILINDRI.MOTOR6[4] := FALSE;
   PartManagmenent.LastPart.NazivniPodatki.CILINDRI.MOTOR6[5] := FALSE;
   PartManagmenent.LastPart.NazivniPodatki.CILINDRI.MOTOR6[6] := FALSE;
   PartManagmenent.LastPart.NazivniPodatki.CILINDRI.MOTOR6[7] := FALSE;
   PartManagmenent.LastPart.NazivniPodatki.CILINDRI.MOTOR6[8] := FALSE;
   PartManagmenent.LastPart.NazivniPodatki.CILINDRI.MOTOR6[9] := FALSE;
   PartManagmenent.LastPart.NazivniPodatki.CILINDRI.MOTOR6[10] := FALSE;
   PartManagmenent.LastPart.NazivniPodatki.CILINDRI.MOTOR6[11] := FALSE;
   PartManagmenent.LastPart.NazivniPodatki.CILINDRI.MOTOR6[12] := FALSE;
   PartManagmenent.LastPart.NazivniPodatki.CILINDRI.MOTOR6[13] := FALSE;
   PartManagmenent.LastPart.NazivniPodatki.CILINDRI.MOTOR6[14] := FALSE;
   PartManagmenent.LastPart.NazivniPodatki.CILINDRI.MOTOR6[15] := FALSE;
   PartManagmenent.LastPart.NazivniPodatki.CILINDRI.MOTOR6[16] := FALSE;
   PartManagmenent.LastPart.NazivniPodatki.CILINDRI.MOTOR6[17] := FALSE;
   PartManagmenent.LastPart.NazivniPodatki.CILINDRI.MOTOR6[18] := FALSE;
   PartManagmenent.LastPart.NazivniPodatki.CILINDRI.MOTOR6[19] := FALSE;
   PartManagmenent.LastPart.NazivniPodatki.CILINDRI.MOTOR6[20] := FALSE;
   PartManagmenent.LastPart.TrenutniPodatki.trenutni_pomik := 100;
   PartManagmenent.LastPart.Oblika.s1[0] := FALSE;
   PartManagmenent.LastPart.Oblika.s1[1] := FALSE;
   PartManagmenent.LastPart.Oblika.s1[2] := FALSE;
   PartManagmenent.LastPart.Oblika.s1[3] := FALSE;
   PartManagmenent.LastPart.Oblika.s1[4] := FALSE;
   PartManagmenent.LastPart.Oblika.s1[5] := FALSE;
   PartManagmenent.LastPart.Oblika.s1[6] := FALSE;
   PartManagmenent.LastPart.Oblika.s1[7] := FALSE;
   PartManagmenent.LastPart.Oblika.s1[8] := FALSE;
   PartManagmenent.LastPart.Oblika.s1[9] := FALSE;
   PartManagmenent.LastPart.Oblika.s1[10] := FALSE;
   PartManagmenent.LastPart.Oblika.s1[11] := FALSE;
   PartManagmenent.LastPart.Oblika.s1[12] := FALSE;
   PartManagmenent.LastPart.Oblika.s1[13] := FALSE;
   PartManagmenent.LastPart.Oblika.s1[14] := FALSE;
   PartManagmenent.LastPart.Oblika.s1[15] := FALSE;
   PartManagmenent.LastPart.Oblika.s1[16] := FALSE;
   PartManagmenent.LastPart.Oblika.s1[17] := FALSE;
   PartManagmenent.LastPart.Oblika.s1[18] := FALSE;
   PartManagmenent.LastPart.Oblika.s1[19] := FALSE;
   PartManagmenent.LastPart.Oblika.s1[20] := FALSE;
   PartManagmenent.LastPart.Oblika.s2[0] := FALSE;
   PartManagmenent.LastPart.Oblika.s2[1] := FALSE;
   PartManagmenent.LastPart.Oblika.s2[2] := FALSE;
   PartManagmenent.LastPart.Oblika.s2[3] := FALSE;
   PartManagmenent.LastPart.Oblika.s2[4] := FALSE;
   PartManagmenent.LastPart.Oblika.s2[5] := FALSE;
   PartManagmenent.LastPart.Oblika.s2[6] := FALSE;
   PartManagmenent.LastPart.Oblika.s2[7] := FALSE;
   PartManagmenent.LastPart.Oblika.s2[8] := FALSE;
   PartManagmenent.LastPart.Oblika.s2[9] := FALSE;
   PartManagmenent.LastPart.Oblika.s2[10] := FALSE;
   PartManagmenent.LastPart.Oblika.s2[11] := FALSE;
   PartManagmenent.LastPart.Oblika.s2[12] := FALSE;
   PartManagmenent.LastPart.Oblika.s2[13] := FALSE;
   PartManagmenent.LastPart.Oblika.s2[14] := FALSE;
   PartManagmenent.LastPart.Oblika.s2[15] := FALSE;
   PartManagmenent.LastPart.Oblika.s2[16] := FALSE;
   PartManagmenent.LastPart.Oblika.s2[17] := FALSE;
   PartManagmenent.LastPart.Oblika.s2[18] := FALSE;
   PartManagmenent.LastPart.Oblika.s2[19] := FALSE;
   PartManagmenent.LastPart.Oblika.s2[20] := FALSE;
   PartManagmenent.PartRecept.NazivniPodatki.SifraIzdelka := 0;
   PartManagmenent.PartRecept.NazivniPodatki.st_pomikov := 8;
   PartManagmenent.PartRecept.NazivniPodatki.st_celic := 8;
   PartManagmenent.PartRecept.NazivniPodatki.st_vrst := 2;
   PartManagmenent.PartRecept.NazivniPodatki.CILINDRI.MOTOR1[1] := FALSE;
   PartManagmenent.PartRecept.NazivniPodatki.CILINDRI.MOTOR1[2] := FALSE;
   PartManagmenent.PartRecept.NazivniPodatki.CILINDRI.MOTOR1[3] := TRUE;
   PartManagmenent.PartRecept.NazivniPodatki.CILINDRI.MOTOR1[4] := FALSE;
   PartManagmenent.PartRecept.NazivniPodatki.CILINDRI.MOTOR1[5] := FALSE;
   PartManagmenent.PartRecept.NazivniPodatki.CILINDRI.MOTOR1[6] := FALSE;
   PartManagmenent.PartRecept.NazivniPodatki.CILINDRI.MOTOR1[7] := FALSE;
   PartManagmenent.PartRecept.NazivniPodatki.CILINDRI.MOTOR1[8] := FALSE;
   PartManagmenent.PartRecept.NazivniPodatki.CILINDRI.MOTOR1[9] := FALSE;
   PartManagmenent.PartRecept.NazivniPodatki.CILINDRI.MOTOR1[10] := FALSE;
   PartManagmenent.PartRecept.NazivniPodatki.CILINDRI.MOTOR1[11] := FALSE;
   PartManagmenent.PartRecept.NazivniPodatki.CILINDRI.MOTOR1[12] := FALSE;
   PartManagmenent.PartRecept.NazivniPodatki.CILINDRI.MOTOR1[13] := FALSE;
   PartManagmenent.PartRecept.NazivniPodatki.CILINDRI.MOTOR1[14] := FALSE;
   PartManagmenent.PartRecept.NazivniPodatki.CILINDRI.MOTOR1[15] := FALSE;
   PartManagmenent.PartRecept.NazivniPodatki.CILINDRI.MOTOR1[16] := FALSE;
   PartManagmenent.PartRecept.NazivniPodatki.CILINDRI.MOTOR1[17] := FALSE;
   PartManagmenent.PartRecept.NazivniPodatki.CILINDRI.MOTOR1[18] := FALSE;
   PartManagmenent.PartRecept.NazivniPodatki.CILINDRI.MOTOR1[19] := FALSE;
   PartManagmenent.PartRecept.NazivniPodatki.CILINDRI.MOTOR1[20] := FALSE;
   PartManagmenent.PartRecept.NazivniPodatki.CILINDRI.MOTOR2[1] := FALSE;
   PartManagmenent.PartRecept.NazivniPodatki.CILINDRI.MOTOR2[2] := FALSE;
   PartManagmenent.PartRecept.NazivniPodatki.CILINDRI.MOTOR2[3] := FALSE;
   PartManagmenent.PartRecept.NazivniPodatki.CILINDRI.MOTOR2[4] := FALSE;
   PartManagmenent.PartRecept.NazivniPodatki.CILINDRI.MOTOR2[5] := FALSE;
   PartManagmenent.PartRecept.NazivniPodatki.CILINDRI.MOTOR2[6] := FALSE;
   PartManagmenent.PartRecept.NazivniPodatki.CILINDRI.MOTOR2[7] := FALSE;
   PartManagmenent.PartRecept.NazivniPodatki.CILINDRI.MOTOR2[8] := FALSE;
   PartManagmenent.PartRecept.NazivniPodatki.CILINDRI.MOTOR2[9] := FALSE;
   PartManagmenent.PartRecept.NazivniPodatki.CILINDRI.MOTOR2[10] := FALSE;
   PartManagmenent.PartRecept.NazivniPodatki.CILINDRI.MOTOR2[11] := FALSE;
   PartManagmenent.PartRecept.NazivniPodatki.CILINDRI.MOTOR2[12] := FALSE;
   PartManagmenent.PartRecept.NazivniPodatki.CILINDRI.MOTOR2[13] := FALSE;
   PartManagmenent.PartRecept.NazivniPodatki.CILINDRI.MOTOR2[14] := FALSE;
   PartManagmenent.PartRecept.NazivniPodatki.CILINDRI.MOTOR2[15] := FALSE;
   PartManagmenent.PartRecept.NazivniPodatki.CILINDRI.MOTOR2[16] := FALSE;
   PartManagmenent.PartRecept.NazivniPodatki.CILINDRI.MOTOR2[17] := FALSE;
   PartManagmenent.PartRecept.NazivniPodatki.CILINDRI.MOTOR2[18] := FALSE;
   PartManagmenent.PartRecept.NazivniPodatki.CILINDRI.MOTOR2[19] := FALSE;
   PartManagmenent.PartRecept.NazivniPodatki.CILINDRI.MOTOR2[20] := FALSE;
   PartManagmenent.PartRecept.NazivniPodatki.CILINDRI.MOTOR3[1] := FALSE;
   PartManagmenent.PartRecept.NazivniPodatki.CILINDRI.MOTOR3[2] := FALSE;
   PartManagmenent.PartRecept.NazivniPodatki.CILINDRI.MOTOR3[3] := FALSE;
   PartManagmenent.PartRecept.NazivniPodatki.CILINDRI.MOTOR3[4] := FALSE;
   PartManagmenent.PartRecept.NazivniPodatki.CILINDRI.MOTOR3[5] := FALSE;
   PartManagmenent.PartRecept.NazivniPodatki.CILINDRI.MOTOR3[6] := FALSE;
   PartManagmenent.PartRecept.NazivniPodatki.CILINDRI.MOTOR3[7] := FALSE;
   PartManagmenent.PartRecept.NazivniPodatki.CILINDRI.MOTOR3[8] := FALSE;
   PartManagmenent.PartRecept.NazivniPodatki.CILINDRI.MOTOR3[9] := FALSE;
   PartManagmenent.PartRecept.NazivniPodatki.CILINDRI.MOTOR3[10] := FALSE;
   PartManagmenent.PartRecept.NazivniPodatki.CILINDRI.MOTOR3[11] := FALSE;
   PartManagmenent.PartRecept.NazivniPodatki.CILINDRI.MOTOR3[12] := FALSE;
   PartManagmenent.PartRecept.NazivniPodatki.CILINDRI.MOTOR3[13] := FALSE;
   PartManagmenent.PartRecept.NazivniPodatki.CILINDRI.MOTOR3[14] := FALSE;
   PartManagmenent.PartRecept.NazivniPodatki.CILINDRI.MOTOR3[15] := FALSE;
   PartManagmenent.PartRecept.NazivniPodatki.CILINDRI.MOTOR3[16] := FALSE;
   PartManagmenent.PartRecept.NazivniPodatki.CILINDRI.MOTOR3[17] := FALSE;
   PartManagmenent.PartRecept.NazivniPodatki.CILINDRI.MOTOR3[18] := FALSE;
   PartManagmenent.PartRecept.NazivniPodatki.CILINDRI.MOTOR3[19] := FALSE;
   PartManagmenent.PartRecept.NazivniPodatki.CILINDRI.MOTOR3[20] := FALSE;
   PartManagmenent.PartRecept.NazivniPodatki.CILINDRI.MOTOR4[1] := FALSE;
   PartManagmenent.PartRecept.NazivniPodatki.CILINDRI.MOTOR4[2] := FALSE;
   PartManagmenent.PartRecept.NazivniPodatki.CILINDRI.MOTOR4[3] := FALSE;
   PartManagmenent.PartRecept.NazivniPodatki.CILINDRI.MOTOR4[4] := FALSE;
   PartManagmenent.PartRecept.NazivniPodatki.CILINDRI.MOTOR4[5] := FALSE;
   PartManagmenent.PartRecept.NazivniPodatki.CILINDRI.MOTOR4[6] := FALSE;
   PartManagmenent.PartRecept.NazivniPodatki.CILINDRI.MOTOR4[7] := FALSE;
   PartManagmenent.PartRecept.NazivniPodatki.CILINDRI.MOTOR4[8] := FALSE;
   PartManagmenent.PartRecept.NazivniPodatki.CILINDRI.MOTOR4[9] := FALSE;
   PartManagmenent.PartRecept.NazivniPodatki.CILINDRI.MOTOR4[10] := FALSE;
   PartManagmenent.PartRecept.NazivniPodatki.CILINDRI.MOTOR4[11] := FALSE;
   PartManagmenent.PartRecept.NazivniPodatki.CILINDRI.MOTOR4[12] := FALSE;
   PartManagmenent.PartRecept.NazivniPodatki.CILINDRI.MOTOR4[13] := FALSE;
   PartManagmenent.PartRecept.NazivniPodatki.CILINDRI.MOTOR4[14] := FALSE;
   PartManagmenent.PartRecept.NazivniPodatki.CILINDRI.MOTOR4[15] := FALSE;
   PartManagmenent.PartRecept.NazivniPodatki.CILINDRI.MOTOR4[16] := FALSE;
   PartManagmenent.PartRecept.NazivniPodatki.CILINDRI.MOTOR4[17] := FALSE;
   PartManagmenent.PartRecept.NazivniPodatki.CILINDRI.MOTOR4[18] := FALSE;
   PartManagmenent.PartRecept.NazivniPodatki.CILINDRI.MOTOR4[19] := FALSE;
   PartManagmenent.PartRecept.NazivniPodatki.CILINDRI.MOTOR4[20] := FALSE;